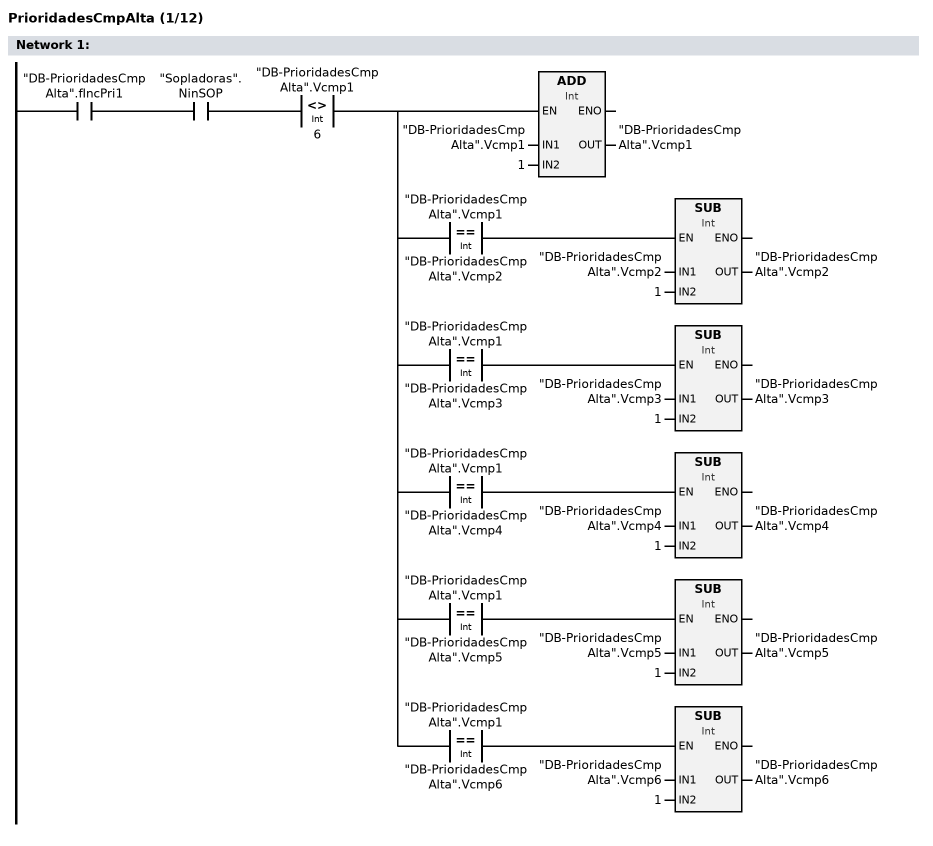
   RUNG wire#powerrail
      Contact( "DB-PrioridadesCmpAlta".fIncPri1 )
      Contact( "Sopladoras".NinSOP )
      { S7_Templates := "SrcType := Int" } NE_Contact(in1 := "DB-PrioridadesCmpAlta".Vcmp1, in2 := 6)
      wire#w1
      { S7_Templates := "SrcType := Int"; S7_GenerateENO := "TRUE" } Add(in1 := "DB-PrioridadesCmpAlta".Vcmp1, in2 := 1, out => "DB-PrioridadesCmpAlta".Vcmp1)
   END_RUNG
   RUNG wire#w1
      { S7_Templates := "SrcType := Int" } EQ_Contact(in1 := "DB-PrioridadesCmpAlta".Vcmp1, in2 := "DB-PrioridadesCmpAlta".Vcmp2)
      { S7_Templates := "SrcType := Int"; S7_GenerateENO := "TRUE" } Sub(in1 := "DB-PrioridadesCmpAlta".Vcmp2, in2 := 1, out => "DB-PrioridadesCmpAlta".Vcmp2)
   END_RUNG
   RUNG wire#w1
      { S7_Templates := "SrcType := Int" } EQ_Contact(in1 := "DB-PrioridadesCmpAlta".Vcmp1, in2 := "DB-PrioridadesCmpAlta".Vcmp3)
      { S7_Templates := "SrcType := Int"; S7_GenerateENO := "TRUE" } Sub(in1 := "DB-PrioridadesCmpAlta".Vcmp3, in2 := 1, out => "DB-PrioridadesCmpAlta".Vcmp3)
   END_RUNG
   RUNG wire#w1
      { S7_Templates := "SrcType := Int" } EQ_Contact(in1 := "DB-PrioridadesCmpAlta".Vcmp1, in2 := "DB-PrioridadesCmpAlta".Vcmp4)
      { S7_Templates := "SrcType := Int"; S7_GenerateENO := "TRUE" } Sub(in1 := "DB-PrioridadesCmpAlta".Vcmp4, in2 := 1, out => "DB-PrioridadesCmpAlta".Vcmp4)
   END_RUNG
   RUNG wire#w1
      { S7_Templates := "SrcType := Int" } EQ_Contact(in1 := "DB-PrioridadesCmpAlta".Vcmp1, in2 := "DB-PrioridadesCmpAlta".Vcmp5)
      { S7_Templates := "SrcType := Int"; S7_GenerateENO := "TRUE" } Sub(in1 := "DB-PrioridadesCmpAlta".Vcmp5, in2 := 1, out => "DB-PrioridadesCmpAlta".Vcmp5)
   END_RUNG
   RUNG wire#w1
      { S7_Templates := "SrcType := Int" } EQ_Contact(in1 := "DB-PrioridadesCmpAlta".Vcmp1, in2 := "DB-PrioridadesCmpAlta".Vcmp6)
      { S7_Templates := "SrcType := Int"; S7_GenerateENO := "TRUE" } Sub(in1 := "DB-PrioridadesCmpAlta".Vcmp6, in2 := 1, out => "DB-PrioridadesCmpAlta".Vcmp6)
   END_RUNG
   // the same network as SCL:
   #_w1 := "DB-PrioridadesCmpAlta".fIncPri1 AND "Sopladoras".NinSOP AND ("DB-PrioridadesCmpAlta".Vcmp1 <> 6);
   IF #_w1 THEN "DB-PrioridadesCmpAlta".Vcmp1 := "DB-PrioridadesCmpAlta".Vcmp1 + 1; END_IF;
   IF #_w1 AND ("DB-PrioridadesCmpAlta".Vcmp1 = "DB-PrioridadesCmpAlta".Vcmp2) THEN
       "DB-PrioridadesCmpAlta".Vcmp2 := "DB-PrioridadesCmpAlta".Vcmp2 - 1;
   END_IF;
   IF #_w1 AND ("DB-PrioridadesCmpAlta".Vcmp1 = "DB-PrioridadesCmpAlta".Vcmp3) THEN
       "DB-PrioridadesCmpAlta".Vcmp3 := "DB-PrioridadesCmpAlta".Vcmp3 - 1;
   END_IF;
   IF #_w1 AND ("DB-PrioridadesCmpAlta".Vcmp1 = "DB-PrioridadesCmpAlta".Vcmp4) THEN
       "DB-PrioridadesCmpAlta".Vcmp4 := "DB-PrioridadesCmpAlta".Vcmp4 - 1;
   END_IF;
   IF #_w1 AND ("DB-PrioridadesCmpAlta".Vcmp1 = "DB-PrioridadesCmpAlta".Vcmp5) THEN
       "DB-PrioridadesCmpAlta".Vcmp5 := "DB-PrioridadesCmpAlta".Vcmp5 - 1;
   END_IF;
   IF #_w1 AND ("DB-PrioridadesCmpAlta".Vcmp1 = "DB-PrioridadesCmpAlta".Vcmp6) THEN
       "DB-PrioridadesCmpAlta".Vcmp6 := "DB-PrioridadesCmpAlta".Vcmp6 - 1;
   END_IF;
END_REGION

REGION Network 2
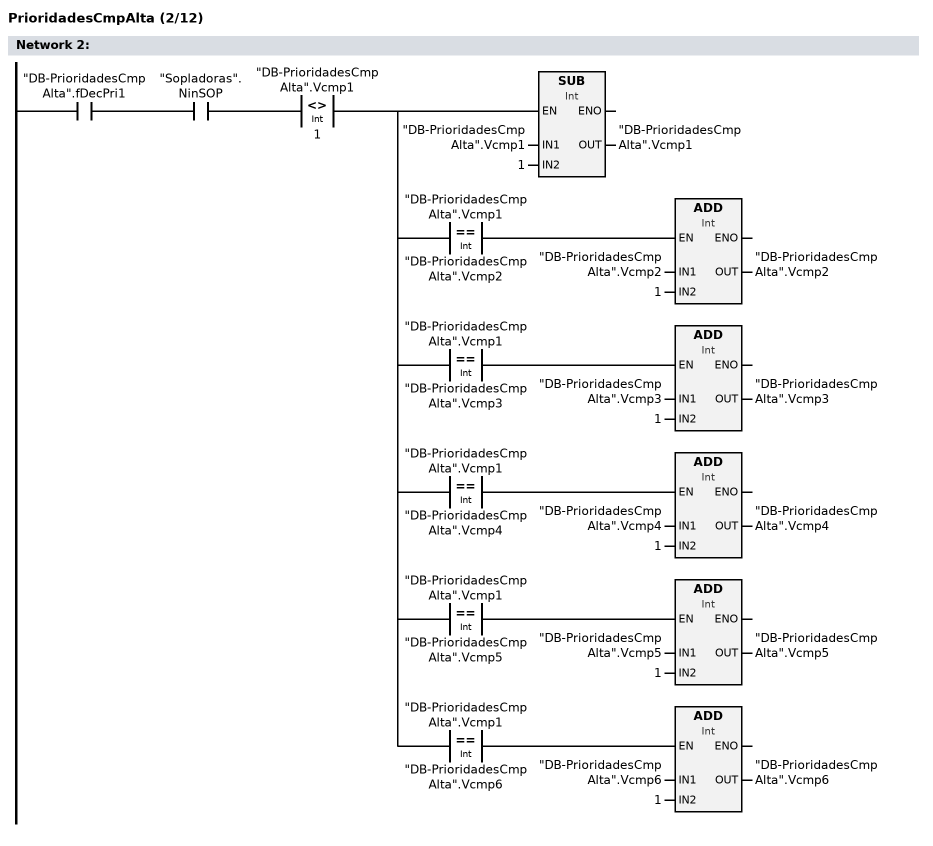
   RUNG wire#powerrail
      Contact( "DB-PrioridadesCmpAlta".fDecPri1 )
      Contact( "Sopladoras".NinSOP )
      { S7_Templates := "SrcType := Int" } NE_Contact(in1 := "DB-PrioridadesCmpAlta".Vcmp1, in2 := 1)
      wire#w1
      { S7_Templates := "SrcType := Int"; S7_GenerateENO := "TRUE" } Sub(in1 := "DB-PrioridadesCmpAlta".Vcmp1, in2 := 1, out => "DB-PrioridadesCmpAlta".Vcmp1)
   END_RUNG
   RUNG wire#w1
      { S7_Templates := "SrcType := Int" } EQ_Contact(in1 := "DB-PrioridadesCmpAlta".Vcmp1, in2 := "DB-PrioridadesCmpAlta".Vcmp2)
      { S7_Templates := "SrcType := Int"; S7_GenerateENO := "TRUE" } Add(in1 := "DB-PrioridadesCmpAlta".Vcmp2, in2 := 1, out => "DB-PrioridadesCmpAlta".Vcmp2)
   END_RUNG
   RUNG wire#w1
      { S7_Templates := "SrcType := Int" } EQ_Contact(in1 := "DB-PrioridadesCmpAlta".Vcmp1, in2 := "DB-PrioridadesCmpAlta".Vcmp3)
      { S7_Templates := "SrcType := Int"; S7_GenerateENO := "TRUE" } Add(in1 := "DB-PrioridadesCmpAlta".Vcmp3, in2 := 1, out => "DB-PrioridadesCmpAlta".Vcmp3)
   END_RUNG
   RUNG wire#w1
      { S7_Templates := "SrcType := Int" } EQ_Contact(in1 := "DB-PrioridadesCmpAlta".Vcmp1, in2 := "DB-PrioridadesCmpAlta".Vcmp4)
      { S7_Templates := "SrcType := Int"; S7_GenerateENO := "TRUE" } Add(in1 := "DB-PrioridadesCmpAlta".Vcmp4, in2 := 1, out => "DB-PrioridadesCmpAlta".Vcmp4)
   END_RUNG
   RUNG wire#w1
      { S7_Templates := "SrcType := Int" } EQ_Contact(in1 := "DB-PrioridadesCmpAlta".Vcmp1, in2 := "DB-PrioridadesCmpAlta".Vcmp5)
      { S7_Templates := "SrcType := Int"; S7_GenerateENO := "TRUE" } Add(in1 := "DB-PrioridadesCmpAlta".Vcmp5, in2 := 1, out => "DB-PrioridadesCmpAlta".Vcmp5)
   END_RUNG
   RUNG wire#w1
      { S7_Templates := "SrcType := Int" } EQ_Contact(in1 := "DB-PrioridadesCmpAlta".Vcmp1, in2 := "DB-PrioridadesCmpAlta".Vcmp6)
      { S7_Templates := "SrcType := Int"; S7_GenerateENO := "TRUE" } Add(in1 := "DB-PrioridadesCmpAlta".Vcmp6, in2 := 1, out => "DB-PrioridadesCmpAlta".Vcmp6)
   END_RUNG
   // the same network as SCL:
   #_w1 := "DB-PrioridadesCmpAlta".fDecPri1 AND "Sopladoras".NinSOP AND ("DB-PrioridadesCmpAlta".Vcmp1 <> 1);
   IF #_w1 THEN "DB-PrioridadesCmpAlta".Vcmp1 := "DB-PrioridadesCmpAlta".Vcmp1 - 1; END_IF;
   IF #_w1 AND ("DB-PrioridadesCmpAlta".Vcmp1 = "DB-PrioridadesCmpAlta".Vcmp2) THEN
       "DB-PrioridadesCmpAlta".Vcmp2 := "DB-PrioridadesCmpAlta".Vcmp2 + 1;
   END_IF;
   IF #_w1 AND ("DB-PrioridadesCmpAlta".Vcmp1 = "DB-PrioridadesCmpAlta".Vcmp3) THEN
       "DB-PrioridadesCmpAlta".Vcmp3 := "DB-PrioridadesCmpAlta".Vcmp3 + 1;
   END_IF;
   IF #_w1 AND ("DB-PrioridadesCmpAlta".Vcmp1 = "DB-PrioridadesCmpAlta".Vcmp4) THEN
       "DB-PrioridadesCmpAlta".Vcmp4 := "DB-PrioridadesCmpAlta".Vcmp4 + 1;
   END_IF;
   IF #_w1 AND ("DB-PrioridadesCmpAlta".Vcmp1 = "DB-PrioridadesCmpAlta".Vcmp5) THEN
       "DB-PrioridadesCmpAlta".Vcmp5 := "DB-PrioridadesCmpAlta".Vcmp5 + 1;
   END_IF;
   IF #_w1 AND ("DB-PrioridadesCmpAlta".Vcmp1 = "DB-PrioridadesCmpAlta".Vcmp6) THEN
       "DB-PrioridadesCmpAlta".Vcmp6 := "DB-PrioridadesCmpAlta".Vcmp6 + 1;
   END_IF;
END_REGION

REGION Network 3
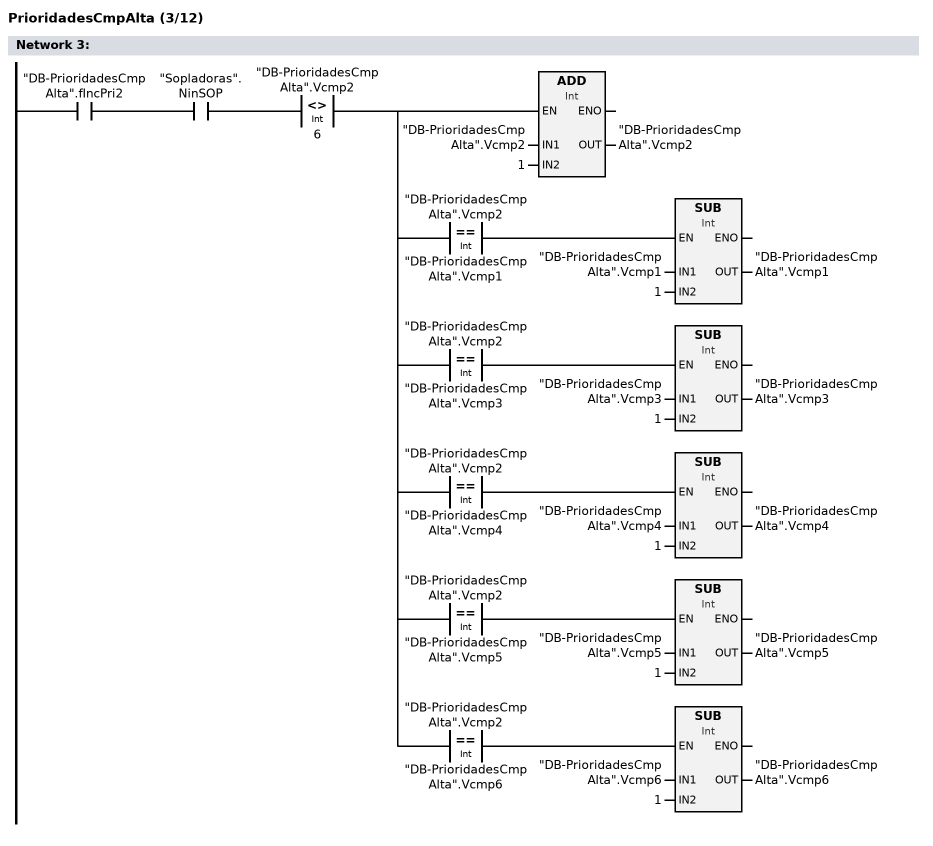
   RUNG wire#powerrail
      Contact( "DB-PrioridadesCmpAlta".fIncPri2 )
      Contact( "Sopladoras".NinSOP )
      { S7_Templates := "SrcType := Int" } NE_Contact(in1 := "DB-PrioridadesCmpAlta".Vcmp2, in2 := 6)
      wire#w1
      { S7_Templates := "SrcType := Int"; S7_GenerateENO := "TRUE" } Add(in1 := "DB-PrioridadesCmpAlta".Vcmp2, in2 := 1, out => "DB-PrioridadesCmpAlta".Vcmp2)
   END_RUNG
   RUNG wire#w1
      { S7_Templates := "SrcType := Int" } EQ_Contact(in1 := "DB-PrioridadesCmpAlta".Vcmp2, in2 := "DB-PrioridadesCmpAlta".Vcmp1)
      { S7_Templates := "SrcType := Int"; S7_GenerateENO := "TRUE" } Sub(in1 := "DB-PrioridadesCmpAlta".Vcmp1, in2 := 1, out => "DB-PrioridadesCmpAlta".Vcmp1)
   END_RUNG
   RUNG wire#w1
      { S7_Templates := "SrcType := Int" } EQ_Contact(in1 := "DB-PrioridadesCmpAlta".Vcmp2, in2 := "DB-PrioridadesCmpAlta".Vcmp3)
      { S7_Templates := "SrcType := Int"; S7_GenerateENO := "TRUE" } Sub(in1 := "DB-PrioridadesCmpAlta".Vcmp3, in2 := 1, out => "DB-PrioridadesCmpAlta".Vcmp3)
   END_RUNG
   RUNG wire#w1
      { S7_Templates := "SrcType := Int" } EQ_Contact(in1 := "DB-PrioridadesCmpAlta".Vcmp2, in2 := "DB-PrioridadesCmpAlta".Vcmp4)
      { S7_Templates := "SrcType := Int"; S7_GenerateENO := "TRUE" } Sub(in1 := "DB-PrioridadesCmpAlta".Vcmp4, in2 := 1, out => "DB-PrioridadesCmpAlta".Vcmp4)
   END_RUNG
   RUNG wire#w1
      { S7_Templates := "SrcType := Int" } EQ_Contact(in1 := "DB-PrioridadesCmpAlta".Vcmp2, in2 := "DB-PrioridadesCmpAlta".Vcmp5)
      { S7_Templates := "SrcType := Int"; S7_GenerateENO := "TRUE" } Sub(in1 := "DB-PrioridadesCmpAlta".Vcmp5, in2 := 1, out => "DB-PrioridadesCmpAlta".Vcmp5)
   END_RUNG
   RUNG wire#w1
      { S7_Templates := "SrcType := Int" } EQ_Contact(in1 := "DB-PrioridadesCmpAlta".Vcmp2, in2 := "DB-PrioridadesCmpAlta".Vcmp6)
      { S7_Templates := "SrcType := Int"; S7_GenerateENO := "TRUE" } Sub(in1 := "DB-PrioridadesCmpAlta".Vcmp6, in2 := 1, out => "DB-PrioridadesCmpAlta".Vcmp6)
   END_RUNG
   // the same network as SCL:
   #_w1 := "DB-PrioridadesCmpAlta".fIncPri2 AND "Sopladoras".NinSOP AND ("DB-PrioridadesCmpAlta".Vcmp2 <> 6);
   IF #_w1 THEN "DB-PrioridadesCmpAlta".Vcmp2 := "DB-PrioridadesCmpAlta".Vcmp2 + 1; END_IF;
   IF #_w1 AND ("DB-PrioridadesCmpAlta".Vcmp2 = "DB-PrioridadesCmpAlta".Vcmp1) THEN
       "DB-PrioridadesCmpAlta".Vcmp1 := "DB-PrioridadesCmpAlta".Vcmp1 - 1;
   END_IF;
   IF #_w1 AND ("DB-PrioridadesCmpAlta".Vcmp2 = "DB-PrioridadesCmpAlta".Vcmp3) THEN
       "DB-PrioridadesCmpAlta".Vcmp3 := "DB-PrioridadesCmpAlta".Vcmp3 - 1;
   END_IF;
   IF #_w1 AND ("DB-PrioridadesCmpAlta".Vcmp2 = "DB-PrioridadesCmpAlta".Vcmp4) THEN
       "DB-PrioridadesCmpAlta".Vcmp4 := "DB-PrioridadesCmpAlta".Vcmp4 - 1;
   END_IF;
   IF #_w1 AND ("DB-PrioridadesCmpAlta".Vcmp2 = "DB-PrioridadesCmpAlta".Vcmp5) THEN
       "DB-PrioridadesCmpAlta".Vcmp5 := "DB-PrioridadesCmpAlta".Vcmp5 - 1;
   END_IF;
   IF #_w1 AND ("DB-PrioridadesCmpAlta".Vcmp2 = "DB-PrioridadesCmpAlta".Vcmp6) THEN
       "DB-PrioridadesCmpAlta".Vcmp6 := "DB-PrioridadesCmpAlta".Vcmp6 - 1;
   END_IF;
END_REGION

REGION Network 4
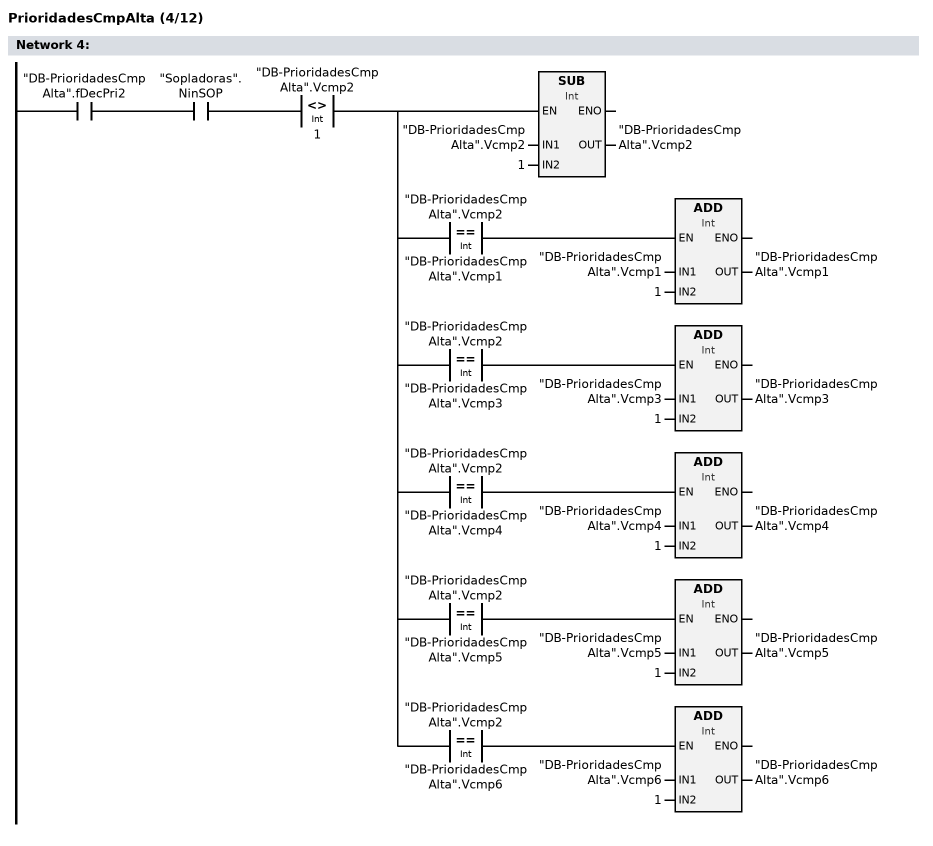
   RUNG wire#powerrail
      Contact( "DB-PrioridadesCmpAlta".fDecPri2 )
      Contact( "Sopladoras".NinSOP )
      { S7_Templates := "SrcType := Int" } NE_Contact(in1 := "DB-PrioridadesCmpAlta".Vcmp2, in2 := 1)
      wire#w1
      { S7_Templates := "SrcType := Int"; S7_GenerateENO := "TRUE" } Sub(in1 := "DB-PrioridadesCmpAlta".Vcmp2, in2 := 1, out => "DB-PrioridadesCmpAlta".Vcmp2)
   END_RUNG
   RUNG wire#w1
      { S7_Templates := "SrcType := Int" } EQ_Contact(in1 := "DB-PrioridadesCmpAlta".Vcmp2, in2 := "DB-PrioridadesCmpAlta".Vcmp1)
      { S7_Templates := "SrcType := Int"; S7_GenerateENO := "TRUE" } Add(in1 := "DB-PrioridadesCmpAlta".Vcmp1, in2 := 1, out => "DB-PrioridadesCmpAlta".Vcmp1)
   END_RUNG
   RUNG wire#w1
      { S7_Templates := "SrcType := Int" } EQ_Contact(in1 := "DB-PrioridadesCmpAlta".Vcmp2, in2 := "DB-PrioridadesCmpAlta".Vcmp3)
      { S7_Templates := "SrcType := Int"; S7_GenerateENO := "TRUE" } Add(in1 := "DB-PrioridadesCmpAlta".Vcmp3, in2 := 1, out => "DB-PrioridadesCmpAlta".Vcmp3)
   END_RUNG
   RUNG wire#w1
      { S7_Templates := "SrcType := Int" } EQ_Contact(in1 := "DB-PrioridadesCmpAlta".Vcmp2, in2 := "DB-PrioridadesCmpAlta".Vcmp4)
      { S7_Templates := "SrcType := Int"; S7_GenerateENO := "TRUE" } Add(in1 := "DB-PrioridadesCmpAlta".Vcmp4, in2 := 1, out => "DB-PrioridadesCmpAlta".Vcmp4)
   END_RUNG
   RUNG wire#w1
      { S7_Templates := "SrcType := Int" } EQ_Contact(in1 := "DB-PrioridadesCmpAlta".Vcmp2, in2 := "DB-PrioridadesCmpAlta".Vcmp5)
      { S7_Templates := "SrcType := Int"; S7_GenerateENO := "TRUE" } Add(in1 := "DB-PrioridadesCmpAlta".Vcmp5, in2 := 1, out => "DB-PrioridadesCmpAlta".Vcmp5)
   END_RUNG
   RUNG wire#w1
      { S7_Templates := "SrcType := Int" } EQ_Contact(in1 := "DB-PrioridadesCmpAlta".Vcmp2, in2 := "DB-PrioridadesCmpAlta".Vcmp6)
      { S7_Templates := "SrcType := Int"; S7_GenerateENO := "TRUE" } Add(in1 := "DB-PrioridadesCmpAlta".Vcmp6, in2 := 1, out => "DB-PrioridadesCmpAlta".Vcmp6)
   END_RUNG
   // the same network as SCL:
   #_w1 := "DB-PrioridadesCmpAlta".fDecPri2 AND "Sopladoras".NinSOP AND ("DB-PrioridadesCmpAlta".Vcmp2 <> 1);
   IF #_w1 THEN "DB-PrioridadesCmpAlta".Vcmp2 := "DB-PrioridadesCmpAlta".Vcmp2 - 1; END_IF;
   IF #_w1 AND ("DB-PrioridadesCmpAlta".Vcmp2 = "DB-PrioridadesCmpAlta".Vcmp1) THEN
       "DB-PrioridadesCmpAlta".Vcmp1 := "DB-PrioridadesCmpAlta".Vcmp1 + 1;
   END_IF;
   IF #_w1 AND ("DB-PrioridadesCmpAlta".Vcmp2 = "DB-PrioridadesCmpAlta".Vcmp3) THEN
       "DB-PrioridadesCmpAlta".Vcmp3 := "DB-PrioridadesCmpAlta".Vcmp3 + 1;
   END_IF;
   IF #_w1 AND ("DB-PrioridadesCmpAlta".Vcmp2 = "DB-PrioridadesCmpAlta".Vcmp4) THEN
       "DB-PrioridadesCmpAlta".Vcmp4 := "DB-PrioridadesCmpAlta".Vcmp4 + 1;
   END_IF;
   IF #_w1 AND ("DB-PrioridadesCmpAlta".Vcmp2 = "DB-PrioridadesCmpAlta".Vcmp5) THEN
       "DB-PrioridadesCmpAlta".Vcmp5 := "DB-PrioridadesCmpAlta".Vcmp5 + 1;
   END_IF;
   IF #_w1 AND ("DB-PrioridadesCmpAlta".Vcmp2 = "DB-PrioridadesCmpAlta".Vcmp6) THEN
       "DB-PrioridadesCmpAlta".Vcmp6 := "DB-PrioridadesCmpAlta".Vcmp6 + 1;
   END_IF;
END_REGION

REGION Network 5
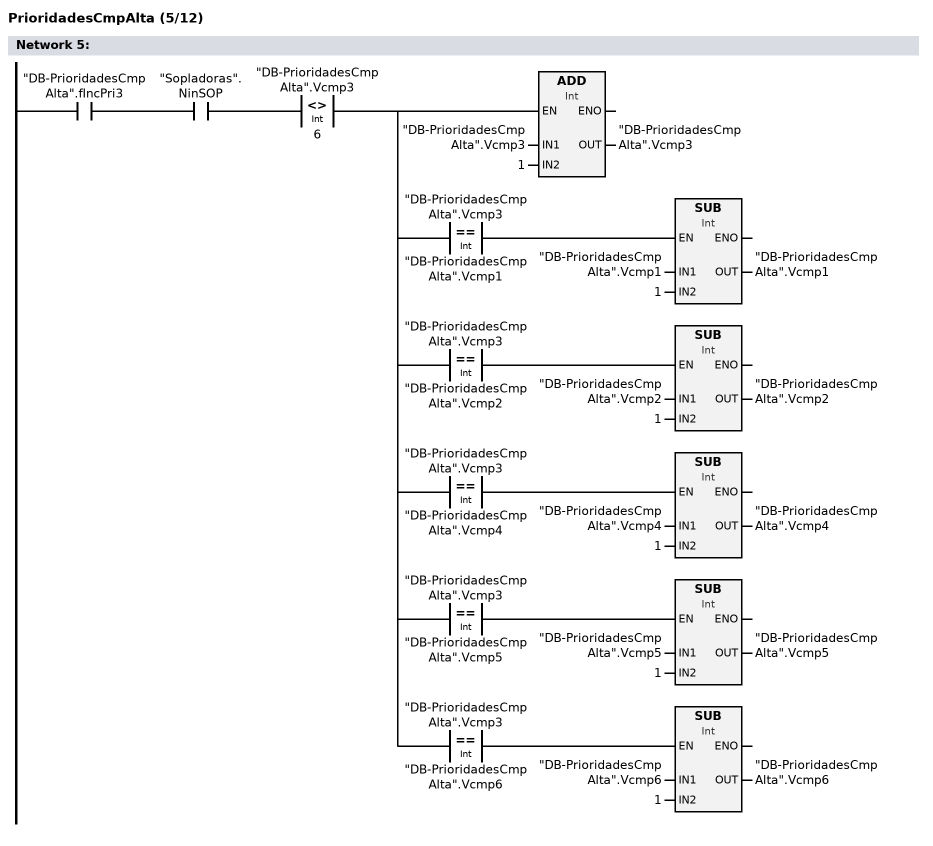
   RUNG wire#powerrail
      Contact( "DB-PrioridadesCmpAlta".fIncPri3 )
      Contact( "Sopladoras".NinSOP )
      { S7_Templates := "SrcType := Int" } NE_Contact(in1 := "DB-PrioridadesCmpAlta".Vcmp3, in2 := 6)
      wire#w1
      { S7_Templates := "SrcType := Int"; S7_GenerateENO := "TRUE" } Add(in1 := "DB-PrioridadesCmpAlta".Vcmp3, in2 := 1, out => "DB-PrioridadesCmpAlta".Vcmp3)
   END_RUNG
   RUNG wire#w1
      { S7_Templates := "SrcType := Int" } EQ_Contact(in1 := "DB-PrioridadesCmpAlta".Vcmp3, in2 := "DB-PrioridadesCmpAlta".Vcmp1)
      { S7_Templates := "SrcType := Int"; S7_GenerateENO := "TRUE" } Sub(in1 := "DB-PrioridadesCmpAlta".Vcmp1, in2 := 1, out => "DB-PrioridadesCmpAlta".Vcmp1)
   END_RUNG
   RUNG wire#w1
      { S7_Templates := "SrcType := Int" } EQ_Contact(in1 := "DB-PrioridadesCmpAlta".Vcmp3, in2 := "DB-PrioridadesCmpAlta".Vcmp2)
      { S7_Templates := "SrcType := Int"; S7_GenerateENO := "TRUE" } Sub(in1 := "DB-PrioridadesCmpAlta".Vcmp2, in2 := 1, out => "DB-PrioridadesCmpAlta".Vcmp2)
   END_RUNG
   RUNG wire#w1
      { S7_Templates := "SrcType := Int" } EQ_Contact(in1 := "DB-PrioridadesCmpAlta".Vcmp3, in2 := "DB-PrioridadesCmpAlta".Vcmp4)
      { S7_Templates := "SrcType := Int"; S7_GenerateENO := "TRUE" } Sub(in1 := "DB-PrioridadesCmpAlta".Vcmp4, in2 := 1, out => "DB-PrioridadesCmpAlta".Vcmp4)
   END_RUNG
   RUNG wire#w1
      { S7_Templates := "SrcType := Int" } EQ_Contact(in1 := "DB-PrioridadesCmpAlta".Vcmp3, in2 := "DB-PrioridadesCmpAlta".Vcmp5)
      { S7_Templates := "SrcType := Int"; S7_GenerateENO := "TRUE" } Sub(in1 := "DB-PrioridadesCmpAlta".Vcmp5, in2 := 1, out => "DB-PrioridadesCmpAlta".Vcmp5)
   END_RUNG
   RUNG wire#w1
      { S7_Templates := "SrcType := Int" } EQ_Contact(in1 := "DB-PrioridadesCmpAlta".Vcmp3, in2 := "DB-PrioridadesCmpAlta".Vcmp6)
      { S7_Templates := "SrcType := Int"; S7_GenerateENO := "TRUE" } Sub(in1 := "DB-PrioridadesCmpAlta".Vcmp6, in2 := 1, out => "DB-PrioridadesCmpAlta".Vcmp6)
   END_RUNG
   // the same network as SCL:
   #_w1 := "DB-PrioridadesCmpAlta".fIncPri3 AND "Sopladoras".NinSOP AND ("DB-PrioridadesCmpAlta".Vcmp3 <> 6);
   IF #_w1 THEN "DB-PrioridadesCmpAlta".Vcmp3 := "DB-PrioridadesCmpAlta".Vcmp3 + 1; END_IF;
   IF #_w1 AND ("DB-PrioridadesCmpAlta".Vcmp3 = "DB-PrioridadesCmpAlta".Vcmp1) THEN
       "DB-PrioridadesCmpAlta".Vcmp1 := "DB-PrioridadesCmpAlta".Vcmp1 - 1;
   END_IF;
   IF #_w1 AND ("DB-PrioridadesCmpAlta".Vcmp3 = "DB-PrioridadesCmpAlta".Vcmp2) THEN
       "DB-PrioridadesCmpAlta".Vcmp2 := "DB-PrioridadesCmpAlta".Vcmp2 - 1;
   END_IF;
   IF #_w1 AND ("DB-PrioridadesCmpAlta".Vcmp3 = "DB-PrioridadesCmpAlta".Vcmp4) THEN
       "DB-PrioridadesCmpAlta".Vcmp4 := "DB-PrioridadesCmpAlta".Vcmp4 - 1;
   END_IF;
   IF #_w1 AND ("DB-PrioridadesCmpAlta".Vcmp3 = "DB-PrioridadesCmpAlta".Vcmp5) THEN
       "DB-PrioridadesCmpAlta".Vcmp5 := "DB-PrioridadesCmpAlta".Vcmp5 - 1;
   END_IF;
   IF #_w1 AND ("DB-PrioridadesCmpAlta".Vcmp3 = "DB-PrioridadesCmpAlta".Vcmp6) THEN
       "DB-PrioridadesCmpAlta".Vcmp6 := "DB-PrioridadesCmpAlta".Vcmp6 - 1;
   END_IF;
END_REGION

REGION Network 6
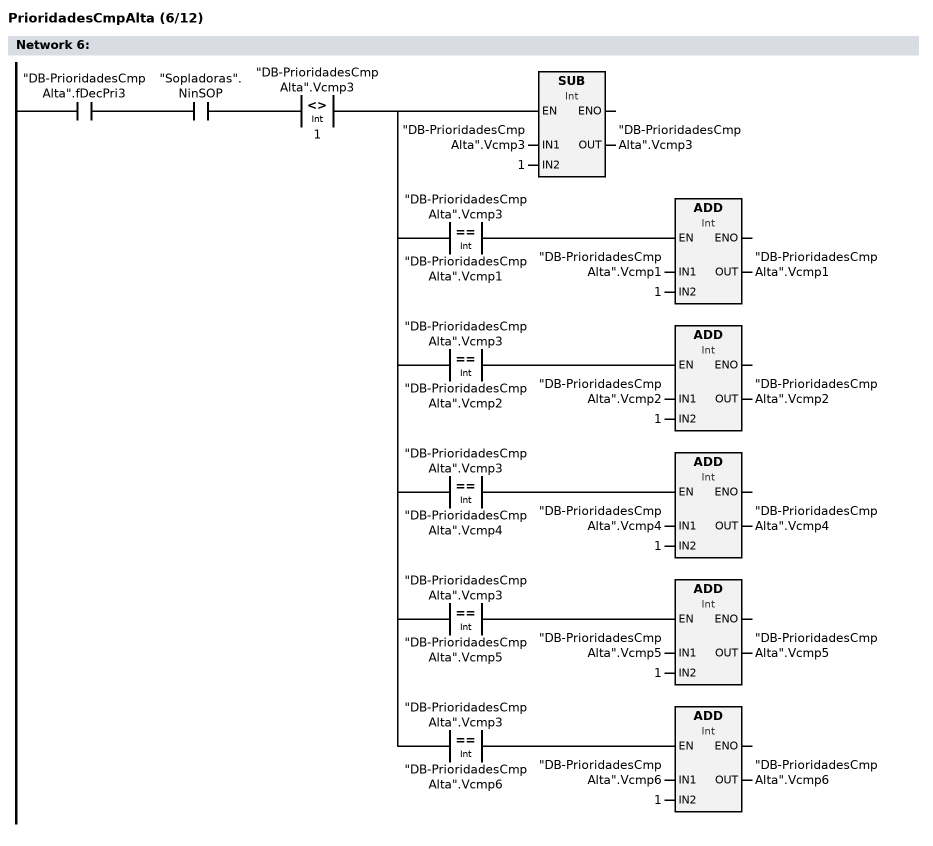
   RUNG wire#powerrail
      Contact( "DB-PrioridadesCmpAlta".fDecPri3 )
      Contact( "Sopladoras".NinSOP )
      { S7_Templates := "SrcType := Int" } NE_Contact(in1 := "DB-PrioridadesCmpAlta".Vcmp3, in2 := 1)
      wire#w1
      { S7_Templates := "SrcType := Int"; S7_GenerateENO := "TRUE" } Sub(in1 := "DB-PrioridadesCmpAlta".Vcmp3, in2 := 1, out => "DB-PrioridadesCmpAlta".Vcmp3)
   END_RUNG
   RUNG wire#w1
      { S7_Templates := "SrcType := Int" } EQ_Contact(in1 := "DB-PrioridadesCmpAlta".Vcmp3, in2 := "DB-PrioridadesCmpAlta".Vcmp1)
      { S7_Templates := "SrcType := Int"; S7_GenerateENO := "TRUE" } Add(in1 := "DB-PrioridadesCmpAlta".Vcmp1, in2 := 1, out => "DB-PrioridadesCmpAlta".Vcmp1)
   END_RUNG
   RUNG wire#w1
      { S7_Templates := "SrcType := Int" } EQ_Contact(in1 := "DB-PrioridadesCmpAlta".Vcmp3, in2 := "DB-PrioridadesCmpAlta".Vcmp2)
      { S7_Templates := "SrcType := Int"; S7_GenerateENO := "TRUE" } Add(in1 := "DB-PrioridadesCmpAlta".Vcmp2, in2 := 1, out => "DB-PrioridadesCmpAlta".Vcmp2)
   END_RUNG
   RUNG wire#w1
      { S7_Templates := "SrcType := Int" } EQ_Contact(in1 := "DB-PrioridadesCmpAlta".Vcmp3, in2 := "DB-PrioridadesCmpAlta".Vcmp4)
      { S7_Templates := "SrcType := Int"; S7_GenerateENO := "TRUE" } Add(in1 := "DB-PrioridadesCmpAlta".Vcmp4, in2 := 1, out => "DB-PrioridadesCmpAlta".Vcmp4)
   END_RUNG
   RUNG wire#w1
      { S7_Templates := "SrcType := Int" } EQ_Contact(in1 := "DB-PrioridadesCmpAlta".Vcmp3, in2 := "DB-PrioridadesCmpAlta".Vcmp5)
      { S7_Templates := "SrcType := Int"; S7_GenerateENO := "TRUE" } Add(in1 := "DB-PrioridadesCmpAlta".Vcmp5, in2 := 1, out => "DB-PrioridadesCmpAlta".Vcmp5)
   END_RUNG
   RUNG wire#w1
      { S7_Templates := "SrcType := Int" } EQ_Contact(in1 := "DB-PrioridadesCmpAlta".Vcmp3, in2 := "DB-PrioridadesCmpAlta".Vcmp6)
      { S7_Templates := "SrcType := Int"; S7_GenerateENO := "TRUE" } Add(in1 := "DB-PrioridadesCmpAlta".Vcmp6, in2 := 1, out => "DB-PrioridadesCmpAlta".Vcmp6)
   END_RUNG
   // the same network as SCL:
   #_w1 := "DB-PrioridadesCmpAlta".fDecPri3 AND "Sopladoras".NinSOP AND ("DB-PrioridadesCmpAlta".Vcmp3 <> 1);
   IF #_w1 THEN "DB-PrioridadesCmpAlta".Vcmp3 := "DB-PrioridadesCmpAlta".Vcmp3 - 1; END_IF;
   IF #_w1 AND ("DB-PrioridadesCmpAlta".Vcmp3 = "DB-PrioridadesCmpAlta".Vcmp1) THEN
       "DB-PrioridadesCmpAlta".Vcmp1 := "DB-PrioridadesCmpAlta".Vcmp1 + 1;
   END_IF;
   IF #_w1 AND ("DB-PrioridadesCmpAlta".Vcmp3 = "DB-PrioridadesCmpAlta".Vcmp2) THEN
       "DB-PrioridadesCmpAlta".Vcmp2 := "DB-PrioridadesCmpAlta".Vcmp2 + 1;
   END_IF;
   IF #_w1 AND ("DB-PrioridadesCmpAlta".Vcmp3 = "DB-PrioridadesCmpAlta".Vcmp4) THEN
       "DB-PrioridadesCmpAlta".Vcmp4 := "DB-PrioridadesCmpAlta".Vcmp4 + 1;
   END_IF;
   IF #_w1 AND ("DB-PrioridadesCmpAlta".Vcmp3 = "DB-PrioridadesCmpAlta".Vcmp5) THEN
       "DB-PrioridadesCmpAlta".Vcmp5 := "DB-PrioridadesCmpAlta".Vcmp5 + 1;
   END_IF;
   IF #_w1 AND ("DB-PrioridadesCmpAlta".Vcmp3 = "DB-PrioridadesCmpAlta".Vcmp6) THEN
       "DB-PrioridadesCmpAlta".Vcmp6 := "DB-PrioridadesCmpAlta".Vcmp6 + 1;
   END_IF;
END_REGION

REGION Network 7
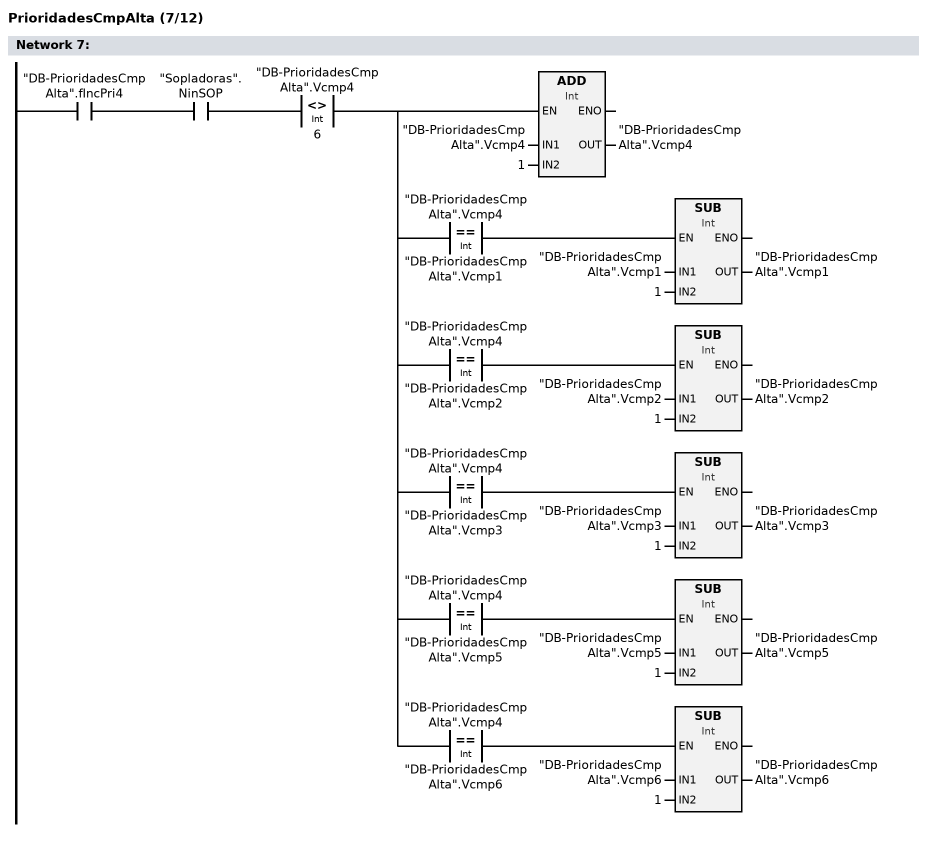
   RUNG wire#powerrail
      Contact( "DB-PrioridadesCmpAlta".fIncPri4 )
      Contact( "Sopladoras".NinSOP )
      { S7_Templates := "SrcType := Int" } NE_Contact(in1 := "DB-PrioridadesCmpAlta".Vcmp4, in2 := 6)
      wire#w1
      { S7_Templates := "SrcType := Int"; S7_GenerateENO := "TRUE" } Add(in1 := "DB-PrioridadesCmpAlta".Vcmp4, in2 := 1, out => "DB-PrioridadesCmpAlta".Vcmp4)
   END_RUNG
   RUNG wire#w1
      { S7_Templates := "SrcType := Int" } EQ_Contact(in1 := "DB-PrioridadesCmpAlta".Vcmp4, in2 := "DB-PrioridadesCmpAlta".Vcmp1)
      { S7_Templates := "SrcType := Int"; S7_GenerateENO := "TRUE" } Sub(in1 := "DB-PrioridadesCmpAlta".Vcmp1, in2 := 1, out => "DB-PrioridadesCmpAlta".Vcmp1)
   END_RUNG
   RUNG wire#w1
      { S7_Templates := "SrcType := Int" } EQ_Contact(in1 := "DB-PrioridadesCmpAlta".Vcmp4, in2 := "DB-PrioridadesCmpAlta".Vcmp2)
      { S7_Templates := "SrcType := Int"; S7_GenerateENO := "TRUE" } Sub(in1 := "DB-PrioridadesCmpAlta".Vcmp2, in2 := 1, out => "DB-PrioridadesCmpAlta".Vcmp2)
   END_RUNG
   RUNG wire#w1
      { S7_Templates := "SrcType := Int" } EQ_Contact(in1 := "DB-PrioridadesCmpAlta".Vcmp4, in2 := "DB-PrioridadesCmpAlta".Vcmp3)
      { S7_Templates := "SrcType := Int"; S7_GenerateENO := "TRUE" } Sub(in1 := "DB-PrioridadesCmpAlta".Vcmp3, in2 := 1, out => "DB-PrioridadesCmpAlta".Vcmp3)
   END_RUNG
   RUNG wire#w1
      { S7_Templates := "SrcType := Int" } EQ_Contact(in1 := "DB-PrioridadesCmpAlta".Vcmp4, in2 := "DB-PrioridadesCmpAlta".Vcmp5)
      { S7_Templates := "SrcType := Int"; S7_GenerateENO := "TRUE" } Sub(in1 := "DB-PrioridadesCmpAlta".Vcmp5, in2 := 1, out => "DB-PrioridadesCmpAlta".Vcmp5)
   END_RUNG
   RUNG wire#w1
      { S7_Templates := "SrcType := Int" } EQ_Contact(in1 := "DB-PrioridadesCmpAlta".Vcmp4, in2 := "DB-PrioridadesCmpAlta".Vcmp6)
      { S7_Templates := "SrcType := Int"; S7_GenerateENO := "TRUE" } Sub(in1 := "DB-PrioridadesCmpAlta".Vcmp6, in2 := 1, out => "DB-PrioridadesCmpAlta".Vcmp6)
   END_RUNG
   // the same network as SCL:
   #_w1 := "DB-PrioridadesCmpAlta".fIncPri4 AND "Sopladoras".NinSOP AND ("DB-PrioridadesCmpAlta".Vcmp4 <> 6);
   IF #_w1 THEN "DB-PrioridadesCmpAlta".Vcmp4 := "DB-PrioridadesCmpAlta".Vcmp4 + 1; END_IF;
   IF #_w1 AND ("DB-PrioridadesCmpAlta".Vcmp4 = "DB-PrioridadesCmpAlta".Vcmp1) THEN
       "DB-PrioridadesCmpAlta".Vcmp1 := "DB-PrioridadesCmpAlta".Vcmp1 - 1;
   END_IF;
   IF #_w1 AND ("DB-PrioridadesCmpAlta".Vcmp4 = "DB-PrioridadesCmpAlta".Vcmp2) THEN
       "DB-PrioridadesCmpAlta".Vcmp2 := "DB-PrioridadesCmpAlta".Vcmp2 - 1;
   END_IF;
   IF #_w1 AND ("DB-PrioridadesCmpAlta".Vcmp4 = "DB-PrioridadesCmpAlta".Vcmp3) THEN
       "DB-PrioridadesCmpAlta".Vcmp3 := "DB-PrioridadesCmpAlta".Vcmp3 - 1;
   END_IF;
   IF #_w1 AND ("DB-PrioridadesCmpAlta".Vcmp4 = "DB-PrioridadesCmpAlta".Vcmp5) THEN
       "DB-PrioridadesCmpAlta".Vcmp5 := "DB-PrioridadesCmpAlta".Vcmp5 - 1;
   END_IF;
   IF #_w1 AND ("DB-PrioridadesCmpAlta".Vcmp4 = "DB-PrioridadesCmpAlta".Vcmp6) THEN
       "DB-PrioridadesCmpAlta".Vcmp6 := "DB-PrioridadesCmpAlta".Vcmp6 - 1;
   END_IF;
END_REGION

REGION Network 8
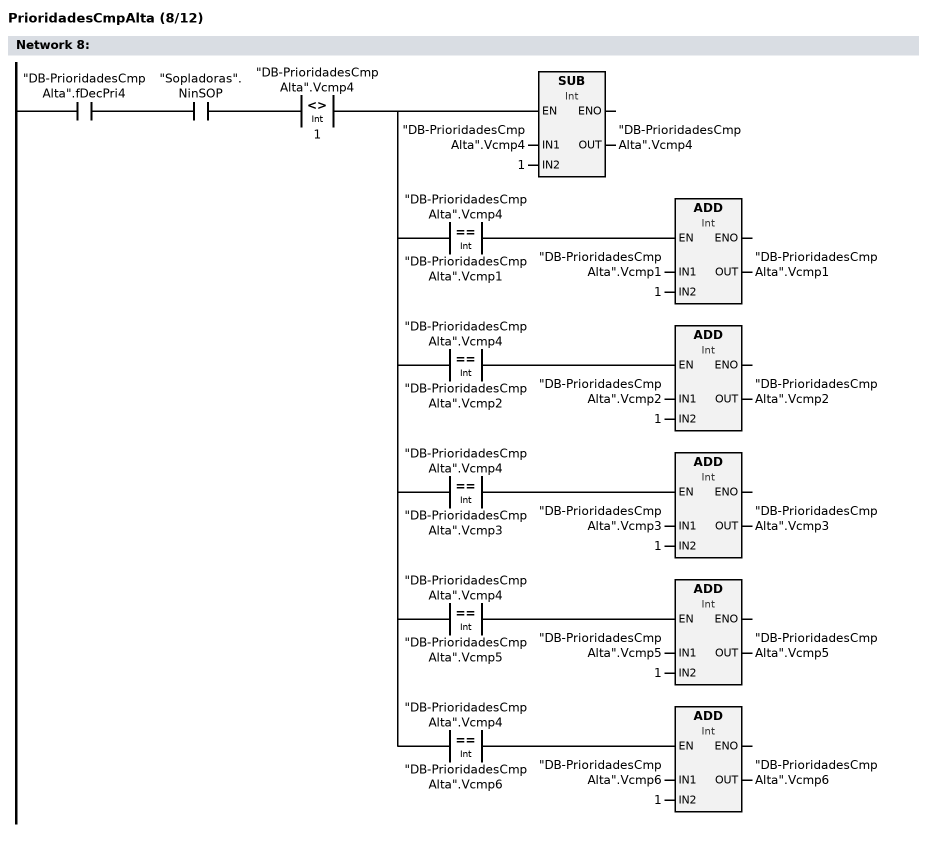
   RUNG wire#powerrail
      Contact( "DB-PrioridadesCmpAlta".fDecPri4 )
      Contact( "Sopladoras".NinSOP )
      { S7_Templates := "SrcType := Int" } NE_Contact(in1 := "DB-PrioridadesCmpAlta".Vcmp4, in2 := 1)
      wire#w1
      { S7_Templates := "SrcType := Int"; S7_GenerateENO := "TRUE" } Sub(in1 := "DB-PrioridadesCmpAlta".Vcmp4, in2 := 1, out => "DB-PrioridadesCmpAlta".Vcmp4)
   END_RUNG
   RUNG wire#w1
      { S7_Templates := "SrcType := Int" } EQ_Contact(in1 := "DB-PrioridadesCmpAlta".Vcmp4, in2 := "DB-PrioridadesCmpAlta".Vcmp1)
      { S7_Templates := "SrcType := Int"; S7_GenerateENO := "TRUE" } Add(in1 := "DB-PrioridadesCmpAlta".Vcmp1, in2 := 1, out => "DB-PrioridadesCmpAlta".Vcmp1)
   END_RUNG
   RUNG wire#w1
      { S7_Templates := "SrcType := Int" } EQ_Contact(in1 := "DB-PrioridadesCmpAlta".Vcmp4, in2 := "DB-PrioridadesCmpAlta".Vcmp2)
      { S7_Templates := "SrcType := Int"; S7_GenerateENO := "TRUE" } Add(in1 := "DB-PrioridadesCmpAlta".Vcmp2, in2 := 1, out => "DB-PrioridadesCmpAlta".Vcmp2)
   END_RUNG
   RUNG wire#w1
      { S7_Templates := "SrcType := Int" } EQ_Contact(in1 := "DB-PrioridadesCmpAlta".Vcmp4, in2 := "DB-PrioridadesCmpAlta".Vcmp3)
      { S7_Templates := "SrcType := Int"; S7_GenerateENO := "TRUE" } Add(in1 := "DB-PrioridadesCmpAlta".Vcmp3, in2 := 1, out => "DB-PrioridadesCmpAlta".Vcmp3)
   END_RUNG
   RUNG wire#w1
      { S7_Templates := "SrcType := Int" } EQ_Contact(in1 := "DB-PrioridadesCmpAlta".Vcmp4, in2 := "DB-PrioridadesCmpAlta".Vcmp5)
      { S7_Templates := "SrcType := Int"; S7_GenerateENO := "TRUE" } Add(in1 := "DB-PrioridadesCmpAlta".Vcmp5, in2 := 1, out => "DB-PrioridadesCmpAlta".Vcmp5)
   END_RUNG
   RUNG wire#w1
      { S7_Templates := "SrcType := Int" } EQ_Contact(in1 := "DB-PrioridadesCmpAlta".Vcmp4, in2 := "DB-PrioridadesCmpAlta".Vcmp6)
      { S7_Templates := "SrcType := Int"; S7_GenerateENO := "TRUE" } Add(in1 := "DB-PrioridadesCmpAlta".Vcmp6, in2 := 1, out => "DB-PrioridadesCmpAlta".Vcmp6)
   END_RUNG
   // the same network as SCL:
   #_w1 := "DB-PrioridadesCmpAlta".fDecPri4 AND "Sopladoras".NinSOP AND ("DB-PrioridadesCmpAlta".Vcmp4 <> 1);
   IF #_w1 THEN "DB-PrioridadesCmpAlta".Vcmp4 := "DB-PrioridadesCmpAlta".Vcmp4 - 1; END_IF;
   IF #_w1 AND ("DB-PrioridadesCmpAlta".Vcmp4 = "DB-PrioridadesCmpAlta".Vcmp1) THEN
       "DB-PrioridadesCmpAlta".Vcmp1 := "DB-PrioridadesCmpAlta".Vcmp1 + 1;
   END_IF;
   IF #_w1 AND ("DB-PrioridadesCmpAlta".Vcmp4 = "DB-PrioridadesCmpAlta".Vcmp2) THEN
       "DB-PrioridadesCmpAlta".Vcmp2 := "DB-PrioridadesCmpAlta".Vcmp2 + 1;
   END_IF;
   IF #_w1 AND ("DB-PrioridadesCmpAlta".Vcmp4 = "DB-PrioridadesCmpAlta".Vcmp3) THEN
       "DB-PrioridadesCmpAlta".Vcmp3 := "DB-PrioridadesCmpAlta".Vcmp3 + 1;
   END_IF;
   IF #_w1 AND ("DB-PrioridadesCmpAlta".Vcmp4 = "DB-PrioridadesCmpAlta".Vcmp5) THEN
       "DB-PrioridadesCmpAlta".Vcmp5 := "DB-PrioridadesCmpAlta".Vcmp5 + 1;
   END_IF;
   IF #_w1 AND ("DB-PrioridadesCmpAlta".Vcmp4 = "DB-PrioridadesCmpAlta".Vcmp6) THEN
       "DB-PrioridadesCmpAlta".Vcmp6 := "DB-PrioridadesCmpAlta".Vcmp6 + 1;
   END_IF;
END_REGION

REGION Network 9
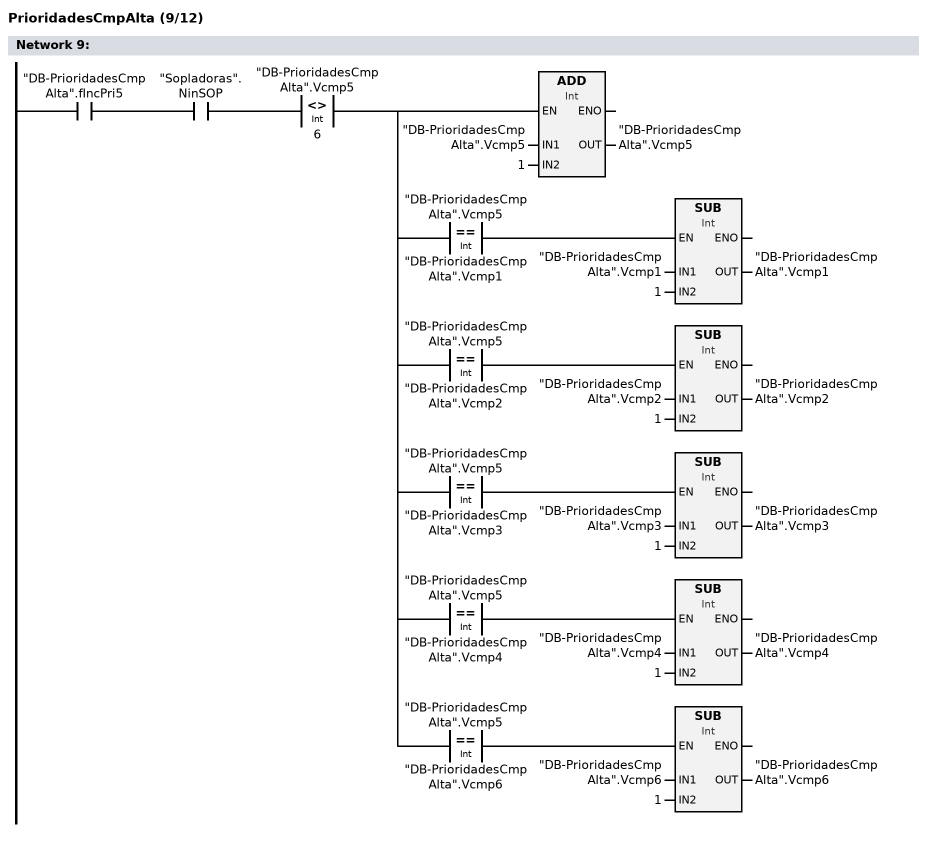
   RUNG wire#powerrail
      Contact( "DB-PrioridadesCmpAlta".fIncPri5 )
      Contact( "Sopladoras".NinSOP )
      { S7_Templates := "SrcType := Int" } NE_Contact(in1 := "DB-PrioridadesCmpAlta".Vcmp5, in2 := 6)
      wire#w1
      { S7_Templates := "SrcType := Int"; S7_GenerateENO := "TRUE" } Add(in1 := "DB-PrioridadesCmpAlta".Vcmp5, in2 := 1, out => "DB-PrioridadesCmpAlta".Vcmp5)
   END_RUNG
   RUNG wire#w1
      { S7_Templates := "SrcType := Int" } EQ_Contact(in1 := "DB-PrioridadesCmpAlta".Vcmp5, in2 := "DB-PrioridadesCmpAlta".Vcmp1)
      { S7_Templates := "SrcType := Int"; S7_GenerateENO := "TRUE" } Sub(in1 := "DB-PrioridadesCmpAlta".Vcmp1, in2 := 1, out => "DB-PrioridadesCmpAlta".Vcmp1)
   END_RUNG
   RUNG wire#w1
      { S7_Templates := "SrcType := Int" } EQ_Contact(in1 := "DB-PrioridadesCmpAlta".Vcmp5, in2 := "DB-PrioridadesCmpAlta".Vcmp2)
      { S7_Templates := "SrcType := Int"; S7_GenerateENO := "TRUE" } Sub(in1 := "DB-PrioridadesCmpAlta".Vcmp2, in2 := 1, out => "DB-PrioridadesCmpAlta".Vcmp2)
   END_RUNG
   RUNG wire#w1
      { S7_Templates := "SrcType := Int" } EQ_Contact(in1 := "DB-PrioridadesCmpAlta".Vcmp5, in2 := "DB-PrioridadesCmpAlta".Vcmp3)
      { S7_Templates := "SrcType := Int"; S7_GenerateENO := "TRUE" } Sub(in1 := "DB-PrioridadesCmpAlta".Vcmp3, in2 := 1, out => "DB-PrioridadesCmpAlta".Vcmp3)
   END_RUNG
   RUNG wire#w1
      { S7_Templates := "SrcType := Int" } EQ_Contact(in1 := "DB-PrioridadesCmpAlta".Vcmp5, in2 := "DB-PrioridadesCmpAlta".Vcmp4)
      { S7_Templates := "SrcType := Int"; S7_GenerateENO := "TRUE" } Sub(in1 := "DB-PrioridadesCmpAlta".Vcmp4, in2 := 1, out => "DB-PrioridadesCmpAlta".Vcmp4)
   END_RUNG
   RUNG wire#w1
      { S7_Templates := "SrcType := Int" } EQ_Contact(in1 := "DB-PrioridadesCmpAlta".Vcmp5, in2 := "DB-PrioridadesCmpAlta".Vcmp6)
      { S7_Templates := "SrcType := Int"; S7_GenerateENO := "TRUE" } Sub(in1 := "DB-PrioridadesCmpAlta".Vcmp6, in2 := 1, out => "DB-PrioridadesCmpAlta".Vcmp6)
   END_RUNG
   // the same network as SCL:
   #_w1 := "DB-PrioridadesCmpAlta".fIncPri5 AND "Sopladoras".NinSOP AND ("DB-PrioridadesCmpAlta".Vcmp5 <> 6);
   IF #_w1 THEN "DB-PrioridadesCmpAlta".Vcmp5 := "DB-PrioridadesCmpAlta".Vcmp5 + 1; END_IF;
   IF #_w1 AND ("DB-PrioridadesCmpAlta".Vcmp5 = "DB-PrioridadesCmpAlta".Vcmp1) THEN
       "DB-PrioridadesCmpAlta".Vcmp1 := "DB-PrioridadesCmpAlta".Vcmp1 - 1;
   END_IF;
   IF #_w1 AND ("DB-PrioridadesCmpAlta".Vcmp5 = "DB-PrioridadesCmpAlta".Vcmp2) THEN
       "DB-PrioridadesCmpAlta".Vcmp2 := "DB-PrioridadesCmpAlta".Vcmp2 - 1;
   END_IF;
   IF #_w1 AND ("DB-PrioridadesCmpAlta".Vcmp5 = "DB-PrioridadesCmpAlta".Vcmp3) THEN
       "DB-PrioridadesCmpAlta".Vcmp3 := "DB-PrioridadesCmpAlta".Vcmp3 - 1;
   END_IF;
   IF #_w1 AND ("DB-PrioridadesCmpAlta".Vcmp5 = "DB-PrioridadesCmpAlta".Vcmp4) THEN
       "DB-PrioridadesCmpAlta".Vcmp4 := "DB-PrioridadesCmpAlta".Vcmp4 - 1;
   END_IF;
   IF #_w1 AND ("DB-PrioridadesCmpAlta".Vcmp5 = "DB-PrioridadesCmpAlta".Vcmp6) THEN